(* Logix 5000 project; controller FV vendor 1 type 14 code 217 rev 31.11; software revision 31.00; part 52 of 63 *)
(* tags used below, declared in another part *)
   Alarm_Reset : BOOL;
   comms_to_blunger_write_enabled : BOOL;
   comms_to_fv_route_write_enabled : BOOL;
   comms_to_mv_route_write_enabled : BOOL;
   CWD : CHECKWORD_FLAGS;
   Default_Check_Time : DINT;
   FR_N10 : INT[265];   // FV_AGING Comms to FV Aging PL C
   FV_B62 : INT[255];   // RESEED FLG
   FV_Comms_from_ct_system : MESSAGE;
   FV_Comms_from_fv_routing_system : MESSAGE;
   FV_Comms_from_mv_routing_system : MESSAGE;
   FV_Comms_from_mv_system : MESSAGE;
   fv_comms_to_blunger : MESSAGE;
   fv_comms_to_blunger_timer : TIMER;
   fv_comms_to_fv_route : MESSAGE;
   fv_comms_to_fv_route_timer : TIMER;
   fv_comms_to_mv_route : MESSAGE;
   fv_comms_to_mv_route_timer : TIMER;
   FV_N13 : INT[255];   // PLC>ME Inter PLC comms traf fic inbound
   FV_N14 : INT[255];   // ME>PLC Inter PLC comms traf fic outbound
   FV_N141 : INT[255];   // YSV1 DATA
   FV_N146 : INT[50];   // FV26, CURRENT FV DATA
   FV_N147 : INT[50];   // FV27, CURRENT FV DATA
   FV_N148 : INT[50];   // FV28, CURRENT FV DATA
   FV_N149 : INT[50];   // FV29, CURRENT FV DATA
   FV_N15 : INT[255];   // COMMS_CTRL Inter PLC comms inte rnal working regs
   FV_N150 : INT[50];   // FV30, CURRENT FV DATA
   FV_N151 : INT[50];   // FV31, CURRENT FV DATA
   FV_N15_63_0_OutputBit : BOOL;
   FV_N15_63_1_OutputBit : BOOL;
   FV_N190 : INT[255];   // MVR COMMS
   FV_N191 : INT[255];   // FVR COMMS
   FV_N60 : INT[255];   // RESEED<PC
   FV_N61 : INT[255];   // RESEED>PC
   FV_N64 : INT[255];   // RESEED_SV
   FV_T16 : TIMER[10];
   FV_T4 : TIMER[10];
   FV_T63 : TIMER[20];
   FV_WYT1R : PlantItem;   // WYT1R
   FV_WYT1R_ALARM : ALARM_DIGITAL;
   FV_WYT1R_D : ALIAS FOR Remote_IO:5:O.Data.14;
   FV_WYT1R_R : ALIAS FOR Remote_IO:7:I.Data.20;
   FV_WYT2R : PlantItem;   // WYT2R
   FV_WYT2R_ALARM : ALARM_DIGITAL;
   FV_WYT2R_D : ALIAS FOR Remote_IO:5:O.Data.15;
   FV_WYT2R_R : ALIAS FOR Remote_IO:7:I.Data.21;
   FV_YSV1R : PlantItem;   // YSV1R
   FV_YSV1R_ALARM : ALARM_DIGITAL;
   FV_YSV1R_D : ALIAS FOR Remote_IO:4:O.Data.10;   // YSV 1 rouser
   FV_YSV1R_R : ALIAS FOR Remote_IO:6:I.Data.12;   // YSV 1 Rouser running f/b
   Item_Faults_Are_Latched : BOOL;
   Item_Simulation_Flag : BOOL;
   MV_Read_YST : MESSAGE;
   MV_Read_YST_TMR : TIMER;
   One_Second_One_Scan : ALIAS FOR One_Second_1_scan;
   reset_msg_interval : BOOL;
   Scada_Pump_Fault_No : DINT;
   Scada_Pump_H_Fault_No : DINT;
   Scada_Pump_T_Fault_No : DINT;
   Unused_Healthy_Feedback : BOOL;
   Unused_NotTripped_Feedback : BOOL;
(* FV_Common, continued *)

ROUTINE FV_PLC_COMMS_7   (* ladder *)
   0: NOP();
   1: XIO(FV_T16[0].DN)TON(FV_T16[0],?,?);
   // Comms with MVSYSTEM
   2: XIC(FV_T16[0].DN)MSG(FV_Comms_from_mv_system);
   // Clear my request to MV system to change last reseeded MV to ageing once acknowledgement received from MV system
   3: XIC(FV_N13[2].0)OSR(FV_N15[63].0,FV_N15_63_0_OutputBit)XIC(FV_N15_63_0_OutputBit)[CLR(FV_N14[1]) ,OTU(FV_N14[2].0) ];
   // Comms with CT System
   4: XIC(FV_T16[0].DN)MSG(FV_Comms_from_ct_system);
   // Clear my request to CT system to change last reseeded CT to ageing once acknowledgement received from CT system
   5: XIC(FV_N13[18].0)OSR(FV_N15[63].1,FV_N15_63_1_OutputBit)XIC(FV_N15_63_1_OutputBit)[CLR(FV_N14[4]) ,OTU(FV_N14[5].0) ];
END_ROUTINE

ROUTINE FV_PLC_COMMS_9   (* ladder *)
   0: XIC(FV_T4[2].DN)XIC(FV_N190[200].1)MSG(FV_Comms_from_mv_routing_system);
   1: COP(FV_N190[0],FV_N190[100],4);
   2: XIC(FV_T4[2].DN)XIC(FV_N191[200].1)COP(FR_N10[100],FV_N191[0],20)AFI()MSG(FV_Comms_from_fv_routing_system);
   3: XIC(FV_N191[0].0)OTE(FV_N191[100].0);
   4: MOV(FV_N146[24],FV_N191[101]);
   5: MOV(FV_N147[24],FV_N191[102]);
   6: MOV(FV_N148[24],FV_N191[103]);
   7: MOV(FV_N149[24],FV_N191[104]);
   8: MOV(FV_N150[24],FV_N191[105]);
   9: MOV(FV_N151[24],FV_N191[106]);
   10: MOV(FV_N191[1],FV_N146[40]);
   11: MOV(FV_N191[2],FV_N147[40]);
   12: MOV(FV_N191[3],FV_N148[40]);
   13: MOV(FV_N191[4],FV_N149[40]);
   14: MOV(FV_N191[5],FV_N150[40]);
   15: MOV(FV_N191[6],FV_N151[40]);
   16: XIO(MV_Read_YST_TMR.DN)TON(MV_Read_YST_TMR,?,?);
   17: XIC(MV_Read_YST_TMR.DN)MSG(MV_Read_YST);
END_ROUTINE

ROUTINE FV_PLC_COMMS_Write_Replacements   (* ladder *)
   // On First Scan Stagger The Write Messages
   0: [XIC(s:fs) ,XIC(reset_msg_interval) OTU(reset_msg_interval) ][MOV(5000,fv_comms_to_fv_route_timer.PRE) MOV(5000,fv_comms_to_mv_route_timer.PRE) MOV(5000,fv_comms_to_blunger_timer.PRE) ,MOV(0,fv_comms_to_fv_route_timer.ACC) MOV(1000,fv_comms_to_mv_route_timer.ACC) MOV(2000,fv_comms_to_blunger_timer.ACC) ];
   // Write Timer To FV Routing
   1: XIO(fv_comms_to_fv_route_timer.DN)TON(fv_comms_to_fv_route_timer,?,?);
   2: XIC(comms_to_fv_route_write_enabled)XIC(fv_comms_to_fv_route_timer.DN)MSG(fv_comms_to_fv_route);
   3: [XIC(fv_comms_to_fv_route.DN) ,XIC(fv_comms_to_fv_route.ER) ]OTU(fv_comms_to_fv_route.DN)OTU(fv_comms_to_fv_route.ER)OTU(fv_comms_to_fv_route.EN);
   // Write Timer To MV Routing
   4: XIO(fv_comms_to_mv_route_timer.DN)TON(fv_comms_to_mv_route_timer,?,?);
   5: XIC(comms_to_mv_route_write_enabled)XIC(fv_comms_to_mv_route_timer.DN)AFI()MSG(fv_comms_to_mv_route);
   6: [XIC(fv_comms_to_mv_route.DN) ,XIC(fv_comms_to_mv_route.ER) ]OTU(fv_comms_to_mv_route.DN)OTU(fv_comms_to_mv_route.ER)OTU(fv_comms_to_mv_route.EN);
   // Write Timer To MV Routing
   7: XIO(fv_comms_to_blunger_timer.DN)TON(fv_comms_to_blunger_timer,?,?);
   8: XIC(comms_to_blunger_write_enabled)XIC(fv_comms_to_blunger_timer.DN)MSG(fv_comms_to_blunger);
   9: [XIC(fv_comms_to_blunger.DN) ,XIC(fv_comms_to_blunger.ER) ]OTU(fv_comms_to_blunger.DN)OTU(fv_comms_to_blunger.ER)OTU(fv_comms_to_blunger.EN);
END_ROUTINE

ROUTINE FV_Pumps   (* ladder *)
   0: [NEQ(FV_YSV1R.DriveBits,0) OTE(FV_YSV1R.CW.[CWD.AUTODRV]) ,[XIC(FV_YSV1R.CW.[CWD.AUTODRV]) XIO(FV_YSV1R.CW.[CWD.MANUAL]) ,XIC(FV_YSV1R.CW.[CWD.MANDRV]) XIC(FV_YSV1R.CW.[CWD.MANUAL]) ] OTE(FV_YSV1R.CW.[CWD.OUTPUT]) ,XIC(FV_YSV1R.CW.[CWD.OUTPUT]) OTE(FV_YSV1R_D) ,XIC(S:FS) [OTU(FV_YSV1R.CW.[CWD.MANUAL]) ,LEQ(FV_YSV1R.CheckTime,0) MOV(Default_Check_Time,FV_YSV1R.CheckTime) ] ,[[XIC(FV_YSV1R_R) XIO(Item_Simulation_Flag) ,XIC(Item_Simulation_Flag) [XIC(FV_YSV1R.CW.[CWD.OUTPUT]) XIO(FV_YSV1R.CW.[CWD.SIMFAIL]) ,XIO(FV_YSV1R.CW.[CWD.OUTPUT]) XIC(FV_YSV1R.CW.[CWD.SIMFAIL]) ] ] OTE(FV_YSV1R.CW.[CWD.RUNFB]) ,[XIC(Item_Simulation_Flag) ,XIC(FV_YSV1R.CW.[CWD.CHECKOFF]) ,XIC(Unused_Healthy_Feedback) ] OTE(FV_YSV1R.CW.[CWD.HEALTHYFB]) ,[XIC(Item_Simulation_Flag) ,XIC(FV_YSV1R.CW.[CWD.CHECKOFF]) ,XIC(Unused_NotTripped_Feedback) ] OTE(FV_YSV1R.CW.[CWD.NOTTRIPPEDFB]) ] ,[XIC(FV_YSV1R.CW.[CWD.OUTPUT]) XIO(FV_YSV1R.CW.[CWD.PREVSCAN]) ,XIO(FV_YSV1R.CW.[CWD.OUTPUT]) XIC(FV_YSV1R.CW.[CWD.PREVSCAN]) ] CLR(FV_YSV1R.CheckTimer) ,XIC(One_Second_One_Scan) LES(FV_YSV1R.CheckTimer,FV_YSV1R.CheckTime) ADD(FV_YSV1R.CheckTimer,1,FV_YSV1R.CheckTimer) ,XIO(FV_YSV1R.CW.[CWD.FAULT]) OTU(FV_YSV1R.CW.[CWD.FAULTLOGGED]) ,[GEQ(FV_YSV1R.CheckTimer,FV_YSV1R.CheckTime) [XIC(FV_YSV1R.CW.[CWD.OUTPUT]) XIO(FV_YSV1R.CW.[CWD.RUNFB]) ,XIO(FV_YSV1R.CW.[CWD.OUTPUT]) XIC(FV_YSV1R.CW.[CWD.RUNFB]) ] ,XIO(FV_YSV1R.CW.[CWD.HEALTHYFB]) ,XIO(FV_YSV1R.CW.[CWD.NOTTRIPPEDFB]) ,XIC(FV_YSV1R.CW.[CWD.FAULT]) XIC(Item_Faults_Are_Latched) ,XIC(FV_YSV1R.CW.[CWD.HIGHLIGHT]) ] XIO(FV_YSV1R.CW.[CWD.CHECKOFF]) XIO(Alarm_Reset) [OTE(FV_YSV1R.CW.[CWD.FAULT]) ,ALMD(FV_YSV1R_ALARM,0,0,0,0) ] ,XIC(FV_YSV1R.CW.[CWD.OUTPUT]) OTE(FV_YSV1R.CW.[CWD.PREVSCAN]) ,XIC(FV_YSV1R.CW.[CWD.FAULT]) EQU(Scada_Pump_Fault_No,0) XIO(FV_YSV1R.CW.[CWD.FAULTLOGGED]) [MOV(20001,Scada_Pump_Fault_No) ,OTL(FV_YSV1R.CW.[CWD.FAULTLOGGED]) ] ,XIO(FV_YSV1R.CW.[CWD.HEALTHYFB]) EQU(Scada_Pump_H_Fault_No,0) XIO(FV_YSV1R.CW.[CWD.HEALTHYFAULTLOGGED]) [MOV(20001,Scada_Pump_H_Fault_No) ,OTL(FV_YSV1R.CW.[CWD.HEALTHYFAULTLOGGED]) ] ,XIO(FV_YSV1R.CW.[CWD.NOTTRIPPEDFB]) EQU(Scada_Pump_H_Fault_No,0) XIO(FV_YSV1R.CW.[CWD.TRIPPEDFAULTLOGGED]) [MOV(20001,Scada_Pump_T_Fault_No) ,OTL(FV_YSV1R.CW.[CWD.TRIPPEDFAULTLOGGED]) ] ];
   1: [NEQ(FV_WYT1R.DriveBits,0) OTE(FV_WYT1R.CW.[CWD.AUTODRV]) ,[XIC(FV_WYT1R.CW.[CWD.AUTODRV]) XIO(FV_WYT1R.CW.[CWD.MANUAL]) ,XIC(FV_WYT1R.CW.[CWD.MANDRV]) XIC(FV_WYT1R.CW.[CWD.MANUAL]) ] OTE(FV_WYT1R.CW.[CWD.OUTPUT]) ,XIC(FV_WYT1R.CW.[CWD.OUTPUT]) OTE(FV_WYT1R_D) ,XIC(S:FS) [OTU(FV_WYT1R.CW.[CWD.MANUAL]) ,LEQ(FV_WYT1R.CheckTime,0) MOV(Default_Check_Time,FV_WYT1R.CheckTime) ] ,[[XIC(FV_WYT1R_R) XIO(Item_Simulation_Flag) ,XIC(Item_Simulation_Flag) [XIC(FV_WYT1R.CW.[CWD.OUTPUT]) XIO(FV_WYT1R.CW.[CWD.SIMFAIL]) ,XIO(FV_WYT1R.CW.[CWD.OUTPUT]) XIC(FV_WYT1R.CW.[CWD.SIMFAIL]) ] ] OTE(FV_WYT1R.CW.[CWD.RUNFB]) ,[XIC(Item_Simulation_Flag) ,XIC(FV_WYT1R.CW.[CWD.CHECKOFF]) ,XIC(Unused_Healthy_Feedback) ] OTE(FV_WYT1R.CW.[CWD.HEALTHYFB]) ,[XIC(Item_Simulation_Flag) ,XIC(FV_WYT1R.CW.[CWD.CHECKOFF]) ,XIC(Unused_NotTripped_Feedback) ] OTE(FV_WYT1R.CW.[CWD.NOTTRIPPEDFB]) ] ,[XIC(FV_WYT1R.CW.[CWD.OUTPUT]) XIO(FV_WYT1R.CW.[CWD.PREVSCAN]) ,XIO(FV_WYT1R.CW.[CWD.OUTPUT]) XIC(FV_WYT1R.CW.[CWD.PREVSCAN]) ] CLR(FV_WYT1R.CheckTimer) ,XIC(One_Second_One_Scan) LES(FV_WYT1R.CheckTimer,FV_WYT1R.CheckTime) ADD(FV_WYT1R.CheckTimer,1,FV_WYT1R.CheckTimer) ,XIO(FV_WYT1R.CW.[CWD.FAULT]) OTU(FV_WYT1R.CW.[CWD.FAULTLOGGED]) ,[GEQ(FV_WYT1R.CheckTimer,FV_WYT1R.CheckTime) [XIC(FV_WYT1R.CW.[CWD.OUTPUT]) XIO(FV_WYT1R.CW.[CWD.RUNFB]) ,XIO(FV_WYT1R.CW.[CWD.OUTPUT]) XIC(FV_WYT1R.CW.[CWD.RUNFB]) ] ,XIO(FV_WYT1R.CW.[CWD.HEALTHYFB]) ,XIO(FV_WYT1R.CW.[CWD.NOTTRIPPEDFB]) ,XIC(FV_WYT1R.CW.[CWD.FAULT]) XIC(Item_Faults_Are_Latched) ,XIC(FV_WYT1R.CW.[CWD.HIGHLIGHT]) ] XIO(FV_WYT1R.CW.[CWD.CHECKOFF]) XIO(Alarm_Reset) [OTE(FV_WYT1R.CW.[CWD.FAULT]) ,ALMD(FV_WYT1R_ALARM,0,0,0,0) ] ,XIC(FV_WYT1R.CW.[CWD.OUTPUT]) OTE(FV_WYT1R.CW.[CWD.PREVSCAN]) ,XIC(FV_WYT1R.CW.[CWD.FAULT]) EQU(Scada_Pump_Fault_No,0) XIO(FV_WYT1R.CW.[CWD.FAULTLOGGED]) [MOV(20001,Scada_Pump_Fault_No) ,OTL(FV_WYT1R.CW.[CWD.FAULTLOGGED]) ] ,XIO(FV_WYT1R.CW.[CWD.HEALTHYFB]) EQU(Scada_Pump_H_Fault_No,0) XIO(FV_WYT1R.CW.[CWD.HEALTHYFAULTLOGGED]) [MOV(20001,Scada_Pump_H_Fault_No) ,OTL(FV_WYT1R.CW.[CWD.HEALTHYFAULTLOGGED]) ] ,XIO(FV_WYT1R.CW.[CWD.NOTTRIPPEDFB]) EQU(Scada_Pump_H_Fault_No,0) XIO(FV_WYT1R.CW.[CWD.TRIPPEDFAULTLOGGED]) [MOV(20001,Scada_Pump_T_Fault_No) ,OTL(FV_WYT1R.CW.[CWD.TRIPPEDFAULTLOGGED]) ] ];
   2: [NEQ(FV_WYT2R.DriveBits,0) OTE(FV_WYT2R.CW.[CWD.AUTODRV]) ,[XIC(FV_WYT2R.CW.[CWD.AUTODRV]) XIO(FV_WYT2R.CW.[CWD.MANUAL]) ,XIC(FV_WYT2R.CW.[CWD.MANDRV]) XIC(FV_WYT2R.CW.[CWD.MANUAL]) ] OTE(FV_WYT2R.CW.[CWD.OUTPUT]) ,XIC(FV_WYT2R.CW.[CWD.OUTPUT]) OTE(FV_WYT2R_D) ,XIC(S:FS) [OTU(FV_WYT2R.CW.[CWD.MANUAL]) ,LEQ(FV_WYT2R.CheckTime,0) MOV(Default_Check_Time,FV_WYT2R.CheckTime) ] ,[[XIC(FV_WYT2R_R) XIO(Item_Simulation_Flag) ,XIC(Item_Simulation_Flag) [XIC(FV_WYT2R.CW.[CWD.OUTPUT]) XIO(FV_WYT2R.CW.[CWD.SIMFAIL]) ,XIO(FV_WYT2R.CW.[CWD.OUTPUT]) XIC(FV_WYT2R.CW.[CWD.SIMFAIL]) ] ] OTE(FV_WYT2R.CW.[CWD.RUNFB]) ,[XIC(Item_Simulation_Flag) ,XIC(FV_WYT2R.CW.[CWD.CHECKOFF]) ,XIC(Unused_Healthy_Feedback) ] OTE(FV_WYT2R.CW.[CWD.HEALTHYFB]) ,[XIC(Item_Simulation_Flag) ,XIC(FV_WYT2R.CW.[CWD.CHECKOFF]) ,XIC(Unused_NotTripped_Feedback) ] OTE(FV_WYT2R.CW.[CWD.NOTTRIPPEDFB]) ] ,[XIC(FV_WYT2R.CW.[CWD.OUTPUT]) XIO(FV_WYT2R.CW.[CWD.PREVSCAN]) ,XIO(FV_WYT2R.CW.[CWD.OUTPUT]) XIC(FV_WYT2R.CW.[CWD.PREVSCAN]) ] CLR(FV_WYT2R.CheckTimer) ,XIC(One_Second_One_Scan) LES(FV_WYT2R.CheckTimer,FV_WYT2R.CheckTime) ADD(FV_WYT2R.CheckTimer,1,FV_WYT2R.CheckTimer) ,XIO(FV_WYT2R.CW.[CWD.FAULT]) OTU(FV_WYT2R.CW.[CWD.FAULTLOGGED]) ,[GEQ(FV_WYT2R.CheckTimer,FV_WYT2R.CheckTime) [XIC(FV_WYT2R.CW.[CWD.OUTPUT]) XIO(FV_WYT2R.CW.[CWD.RUNFB]) ,XIO(FV_WYT2R.CW.[CWD.OUTPUT]) XIC(FV_WYT2R.CW.[CWD.RUNFB]) ] ,XIO(FV_WYT2R.CW.[CWD.HEALTHYFB]) ,XIO(FV_WYT2R.CW.[CWD.NOTTRIPPEDFB]) ,XIC(FV_WYT2R.CW.[CWD.FAULT]) XIC(Item_Faults_Are_Latched) ,XIC(FV_WYT2R.CW.[CWD.HIGHLIGHT]) ] XIO(FV_WYT2R.CW.[CWD.CHECKOFF]) XIO(Alarm_Reset) [OTE(FV_WYT2R.CW.[CWD.FAULT]) ,ALMD(FV_WYT2R_ALARM,0,0,0,0) ] ,XIC(FV_WYT2R.CW.[CWD.OUTPUT]) OTE(FV_WYT2R.CW.[CWD.PREVSCAN]) ,XIC(FV_WYT2R.CW.[CWD.FAULT]) EQU(Scada_Pump_Fault_No,0) XIO(FV_WYT2R.CW.[CWD.FAULTLOGGED]) [MOV(20001,Scada_Pump_Fault_No) ,OTL(FV_WYT2R.CW.[CWD.FAULTLOGGED]) ] ,XIO(FV_WYT2R.CW.[CWD.HEALTHYFB]) EQU(Scada_Pump_H_Fault_No,0) XIO(FV_WYT2R.CW.[CWD.HEALTHYFAULTLOGGED]) [MOV(20001,Scada_Pump_H_Fault_No) ,OTL(FV_WYT2R.CW.[CWD.HEALTHYFAULTLOGGED]) ] ,XIO(FV_WYT2R.CW.[CWD.NOTTRIPPEDFB]) EQU(Scada_Pump_H_Fault_No,0) XIO(FV_WYT2R.CW.[CWD.TRIPPEDFAULTLOGGED]) [MOV(20001,Scada_Pump_T_Fault_No) ,OTL(FV_WYT2R.CW.[CWD.TRIPPEDFAULTLOGGED]) ] ];
END_ROUTINE

ROUTINE FV_RESEED_CP_31   (* ladder *)
   // Reset command interpreter step counter
   0: XIC(S:FS)CLR(FV_N61[16]);
   // RESET
   1: EQU(FV_N61[16],0)MCR();
   2: OTU(FV_B62[0].0);
   3: OTU(FV_B62[0].1);
   4: OTU(FV_B62[0].8);
   5: FLL(0,FV_N61[0],16);
   // Set PCparameter buffer to 'Null' value
   6: FLL(-32768,FV_N60[1],7);
   7: CLR(FV_N60[0]);
   8: MOV(1,FV_N61[16]);
   9: MCR();
   // ALLOW STARTUP DIALOG
   10: EQU(FV_N61[16],1)MCR();
   // Set process status = ready
   11: MOV(1,FV_N61[0]);
   // Allow startup if YSV1 is inactive or on storage control only and reseeding line is clean
   12: [EQU(FV_N141[0],0) ,EQU(FV_N141[0],5) ]OTE(FV_N61[2].0);
   // Advance step if start selected
   13: XIC(FV_N61[2].0)XIC(FV_N60[0].0)MOV(2,FV_N61[16]);
   14: MCR();
   // WAIT FOR STARTUP DIALOG COMPLETE
   15: EQU(FV_N61[16],2)MCR();
   // If YSV1 requested and YSV1 not involved in any other startup dialog set lock flag
   // Used to Allow within PLC Startup if 0 , Now disabled to match what it locks out in PC.
   16: EQU(FV_N60[1],1)[EQU(FV_N141[0],0) ,EQU(FV_N141[0],5) ][EQU(FV_N141[4],0) ,XIC(FV_N141[4].5) ]OTE(FV_N141[4].5);
   // Allow start confirmed button if selected YSV could be locked
   17: XIC(FV_N141[4].5)OTE(FV_N61[2].1);
   // Startup dialog guard timer
   18: TON(FV_T63[0],?,?);
   // Reset command processor if dialog cancel selected or startup dialog timer expired
   19: [XIC(FV_N60[0].15) ,XIC(FV_T63[0].DN) ]CLR(FV_N61[16]);
   // Advance step if start available and selected
   20: XIC(FV_N60[0].1)XIC(FV_N61[2].1)[MOV(3,FV_N61[16]) ,CLR(FV_N60[0]) ];
   21: MCR();
   // COMPLETE STARTUP DIALOG
   22: EQU(FV_N61[16],3)MCR();
   // set YSV1 status = Reseeding
   23: EQU(FV_N60[1],1)MOV(6,FV_N141[0]);
   // Set YSV Reseeding Process Status = Running
   24: MOV(2,FV_N61[0]);
   25: OTL(FV_B62[0].0);
   26: OTL(FV_B62[0].1);
   27: OTL(FV_N61[2].2);
   28: MOV(10,FV_N61[1]);
   29: MOV(10,FV_N61[3]);
   30: MOV(-1,FV_N61[16]);
   31: CLR(FV_N60[0]);
   32: MCR();
   // HANDLE STOP BUTTON
   33: XIC(FV_N60[0].2)XIC(FV_N61[2].2)MCR();
   34: OTU(FV_B62[0].1);
   35: OTU(FV_N61[2].2);
   36: OTL(FV_N61[2].3);
   37: OTL(FV_N61[2].4);
   38: MOV(3,FV_N61[0]);
   39: MOV(0,FV_N61[1]);
   40: CLR(FV_N60[0]);
   41: MCR();
   // HANDLE CONTINUE BUTTON
   42: XIC(FV_N60[0].3)XIC(FV_N61[2].3)MCR();
   43: OTL(FV_B62[0].1);
   44: OTL(FV_N61[2].2);
   45: OTU(FV_N61[2].3);
   // Reset process alarm and parameters
   46: OTU(FV_N61[2].4);
   47: FLL(0,FV_N61[4],4);
   48: MOV(2,FV_N61[0]);
   // Set current Step = Restart Step
   49: MOV(FV_N61[3],FV_N61[1]);
   50: CLR(FV_N60[0]);
   51: MCR();
   // HANDLE ABORT BUTTON
   52: XIC(FV_N60[0].4)XIC(FV_N61[2].4)MCR();
   53: OTU(FV_B62[0].0);
   // Set YSV's operation to storage
   54: JSR(FV_Set_FV_Datafile_Value,3,5,FV_N61[15],0);
   55: JSR(FV_Set_FV_Datafile_Value,3,0,FV_N61[15],3);
   56: [MOV(FV_N60[1],FV_N64[1]) ,MOV(FV_N61[10],FV_N64[2]) ,MOV(FV_N60[3],FV_N64[3]) ,MOV(FV_N60[4],FV_N64[4]) ,OTL(FV_N64[0].0) ];
   // Send MV number which was reseeded to MV attemporation system so it can set control to ageing
   57: [LIM(29,FV_N60[4],56) ,EQU(FV_N60[4],94) ,LIM(336,FV_N60[4],347) ][MOV(FV_N60[4],FV_N14[1]) ,OTL(FV_N14[2].0) ];
   // Send CT number which was reseeded to CT attemporation system so it can set control to conditioning
   58: LIM(57,FV_N60[4],91)[MOV(FV_N60[4],FV_N14[4]) ,OTL(FV_N14[5].0) ];
   59: CLR(FV_N61[16]);
   60: CLR(FV_N60[0]);
   61: MCR();
   // Copy step number for PC to display if running
   62: XIC(FV_B62[0].1)MOV(FV_N61[1],FV_N61[9]);
END_ROUTINE
